// TIA Portal project "NX_PLC_Project" (V16)

(* hardware
DEVICE "S71500/ET200MP station_1"  S7-1500 station
   slot 0: "Rail_0"  Rack  6ES7 590-1***0-0AA0
   slot 0: "PM 190W 120/230VAC"  PM 190W 120/230VAC  6EP1333-4BA00
   slot 1: "PLC_1"  CPU 1516-3 PN/DP  6ES7 516-3AN01-0AB0  V2.8
      slot 3: "CPU display_1"  6ES7591-1BA00-0AA0
      slot 32768: "PROFINET interface_1"  X1
         slot 32769: "Port_1"  X1 P1
         slot 32770: "Port_2"  X1 P2
      slot 33024: "PROFINET interface_2"  X2
         slot 33025: "Port_1"  X2 P1
      slot 33280: "DP interface_1"  X3
      slot 34817: "Virtual CP interface port_1"  Virtual CP interface port  Virtual CP interface port
   slot 2: "DI 32x24VDC HF_1"  DI 32x24VDC HF  6ES7 521-1BL00-0AB0  V2.0
   slot 3: "DQ 32x24VDC/0.5A HF_1"  DQ 32x24VDC/0.5A HF  6ES7 522-1BL01-0AB0  V1.0
DEVICE "PC station"  SIMATIC PC station
   slot 0: "PC station"  Rail  SIMATIC PC-Station  V1.0
      slot 125: "Stationmanager"  Station_Manager  V6.0.4
   slot 1: "IE general_1"  IE General  IE_CP  V8.2.0
   slot 2: "HMI_RT_1"  WinCC RT Advanced  6AV2 104-0xxxx-xxxx  16.0.0.0
      slot 33792: "Computer interface"  Host interface
DEVICE "S71500/ET200MP station_2"  S7-1500 station
   slot 0: "Rail_0"  Rack  6ES7 590-1***0-0AA0
   slot 0: "PM 190W 120/230VAC"  PM 190W 120/230VAC  6EP1333-4BA00
   slot 1: "PLC_2"  CPU 1516-3 PN/DP  6ES7 516-3AN01-0AB0  V2.8
      slot 3: "CPU display_1"  6ES7591-1BA00-0AA0
      slot 32768: "PROFINET interface_1"  X1
         slot 32769: "Port_1"  X1 P1
         slot 32770: "Port_2"  X1 P2
      slot 33024: "PROFINET interface_2"  X2
         slot 33025: "Port_1"  X2 P1
      slot 33280: "DP interface_1"  X3
      slot 34817: "Virtual CP interface port_1"  Virtual CP interface port  Virtual CP interface port
   slot 2: "DI 32x24VDC HF_1"  DI 32x24VDC HF  6ES7 521-1BL00-0AB0  V2.0
   slot 3: "DQ 32x24VDC/0.5A HF_1"  DQ 32x24VDC/0.5A HF  6ES7 522-1BL01-0AB0  V1.0
DEVICE "HMI_1"  KTP700 Basic PN
   slot 0: "HMI_1"  KTP700 Basic PN  6AV2 123-2GB03-0AX0  16.0.0.0
   slot 1: "HMI_RT_2"  KTP700 Basic PN  6AV2 123-2GB03-0AX0  16.0.0.0
   slot 5: "HMI_1.IE_CP_1"  PROFINET Interface  16.0.0.0
      slot 1: "PROFINET Interface_1"  PROFINET Interface
         slot 1: "Port_1"  Port
*)

// ===== PLC "PLC_1"  CPU 1516-3 PN/DP =====

VAR_GLOBAL   // PLC tag table "Default tag table"
   "sensor1" AT %I0.0 : Bool;
   "belt1" AT %Q2.0 : Bool;
   "ABB1_ON" AT %M1.3 : Bool;
   "sensor2" AT %I0.1 : Bool;
   "sensor3" AT %I0.3 : Bool;
   "sensor4" AT %I0.4 : Bool;
   "belt2_1" AT %Q0.1 : Bool;
   "belt2_2" AT %Q0.2 : Bool;
   "belt2_3" AT %Q0.3 : Bool;
   "belt3" AT %Q0.4 : Bool;
   "send_small" AT %Q1.1 : Bool;
   "sensor2_tall" AT %I0.2 : Bool;
   "ABB2_IDLE" AT %M1.4 : Bool;
   "send_tall" AT %Q1.0 : Bool;
   "ABB2_ON" AT %M1.5 : Bool;
   "F_IDLE" AT %M0.0 : Bool;
   "FILL_TIMER_COUNT" AT %MD2 : Time;
   "ABB1_IDLE" AT %M1.2 : Bool;
   "F_SEND" AT %M0.1 : Bool;
   "robot1_end" AT %I1.1 : Bool;
   "sensor4_tall" AT %I0.5 : Bool;
   "new_cap" AT %Q1.2 : Bool;
   "F_FILL" AT %M0.2 : Bool;
   "sensor5" AT %I0.6 : Bool;
   "sensor5_tall" AT %I0.7 : Bool;
   "robot1_place_tall" AT %Q1.4 : Bool;
   "robot2_get_tall" AT %Q1.6 : Bool;
   "robot1_place_short" AT %Q1.5 : Bool;
   "robot2_get_short" AT %Q1.7 : Bool;
   "robot2_end" AT %I1.2 : Bool;
   "belt_F" AT %Q0.5 : Bool;
   "belt_L" AT %Q0.6 : Bool;
   "belt_R" AT %Q0.7 : Bool;
   "robot1_getCap" AT %Q1.3 : Bool;
   "Connect" AT %M2.0 : Bool;
   "Send" AT %M2.1 : Bool;
   "Clock_10Hz" AT %M100.0 : Bool;
   "sensor_T" AT %I2.1 : Bool;
   "ABB1_MODE" AT %M1.6 : Bool;
   "ABB2_MODE" AT %M1.7 : Bool;
   "sensor_S" AT %I2.2 : Bool;
   "ABB1_SEND" AT %M6.0 : Bool;
   "robot1_hasCap" AT %I1.0 : Bool;
   "SB_WAIT" AT %M0.3 : Bool;
   "SB_SEND" AT %M0.4 : Bool;
   "CONTROL_ENABLE" AT %M0.5 : Bool;
   "F_RELEASE" AT %M0.6 : Bool;
   "START" AT %I100.0 : Bool;
   "STOP" AT %I100.1 : Bool;
   "RESET" AT %I100.2 : Bool;
   "sink" AT %Q100.3 : Bool;
   "RESTARTING" AT %M0.7 : Bool;
   "ABB1_GETCAP" AT %M1.0 : Bool;
   "END_RESTART" AT %M1.1 : Bool;
END_VAR

DATA_BLOCK "Data_block_1"   // DB3
{ S7_Optimized_Access := 'TRUE' }
VERSION : 0.1
   VAR
      Received_string : String;
      Sent_string : String := 'Hello PLC2';
      Received_array : Array[0..1] of Char;
      Sent_array : Array[0..1] of Char;
   END_VAR
BEGIN
END_DATA_BLOCK

// folder: System blocks/Program resources

DATA_BLOCK "FILL_TIMER"   // DB1
{ S7_Optimized_Access := 'TRUE' }
AUTHOR : Simatic
FAMILY : IEC
NAME : IEC_TMR
VERSION : 1.0
// stored: InstanceOfName IEC_TIMER
"IEC_TIMER"
BEGIN
END_DATA_BLOCK

DATA_BLOCK "sink_timer"   // DB4
{ S7_Optimized_Access := 'TRUE' }
AUTHOR : Simatic
FAMILY : IEC
NAME : IEC_TMR
VERSION : 1.0
// stored: InstanceOfName IEC_TIMER
"IEC_TIMER"
BEGIN
END_DATA_BLOCK

DATA_BLOCK "PLC_1_Connection_DB"   // DB5
{ S7_Optimized_Access := 'TRUE' }
AUTHOR : SIMATIC
FAMILY : MC7Plus
NAME : TC_IP_v4
VERSION : 1.0
// stored: InstanceOfName TCON_IP_v4
"TCON_IP_v4"
BEGIN
   ID := 1;
   InterfaceId := 64;
   LocalPort := 2000;
   RemoteAddress.ADDR[1] := 192;
   RemoteAddress.ADDR[2] := 168;
   RemoteAddress.ADDR[4] := 2;
END_DATA_BLOCK

// folder: (top level)

ORGANIZATION_BLOCK "Main"   // OB1, LAD, ProgramCycle
TITLE = LADDER CODE FOR NX SIMULATION OF WATER BOTTLE ASSEMBLY LINE
{ S7_Optimized_Access := 'TRUE' }
VERSION : 0.1
// This program provides the control logic for an NX simulation via TIA Portal and PLCSIM. The simulation emulates a streamlined factory bottling line where bottles are filled, capped, and sorted for packing based on their size. The production line is organized into two primary stations:
// 
// STATION 1: Filling and Capping. This station processes the initial bottle, which is introduced from an external source (triggered via the HMI). The process begins with filling, where the bottle is conveyed to a valve and held in place for a simulated duration. Once filled, the bottle advances to the working area of ABB Robot 1. Upon detecting the bottle, the robot applies a cap and releases it toward the next stage of the line.
// 
// STATION 2: Sorting and Packing. The second station is responsible for sorting bottles by size to ensure they are packed correctly. When a bottle enters the workspace of ABB Robot 2, the robot identifies its dimensions and, following instructions from the PLC, transfers it to the appropriate secondary conveyor. Finally, the bottle travels down the designated belt to its corresponding packing crate.
// 
// IMPORTANT: The PLC program is architected using three distinct Finite State Machines (FSMs). This modular approach ensures that the Filling, Capping, and Sorting sequences operate independently yet in perfect synchronization. Without this modularity, if we used a single FSM, then instead of having mulltiple bottles going through the process, we would just be tracking a single bottle at a time and this is extremely inefficient. Having this modular approach allows us to only care about the bottles that are going through each process, not the ones moving through the belt.
// 
// IMPORTANT: Even though there are three distinct FSMs, they are connected by the sensors and the input received from the PLC's HMI, which allows us to Start, Stop, and Reset the process at any time. (We can also track the states of the robots and belts)
   VAR_INPUT
      Initial_Call : Bool;   // Initial call of this OB
      Remanence : Bool;   // =True, if remanent data are available
   END_VAR
   VAR_TEMP
      COUNT1 : Int;
      SEND_TIMER_COUNT : Time;
      cnt : UInt;
   END_VAR
   VAR_TEMP   // added for the SCL form of the ladder/FBD networks
      _w1 : Bool;
      _w2 : Bool;
      _w3 : Bool;
      _w4 : Bool;
      _w5 : Bool;
   END_VAR
BEGIN

REGION Network 1: START AND STOP LOGIC
   // This network corresponds to the START and STOP buttons in the HMI. The logic is simple: 
   // 
   // - Branch 1: If the START button is pressed, then the system (CONTROL_ENABLE) is activated.
   // 
   // - Branch 2: If the STOP button is pressed, then the system is turned off.
   // 
   // - Branch 3: If the system (CONTROL_ENABLE) is on, then belt 2 is active (belt 2 is composed of three small belts due to curving)
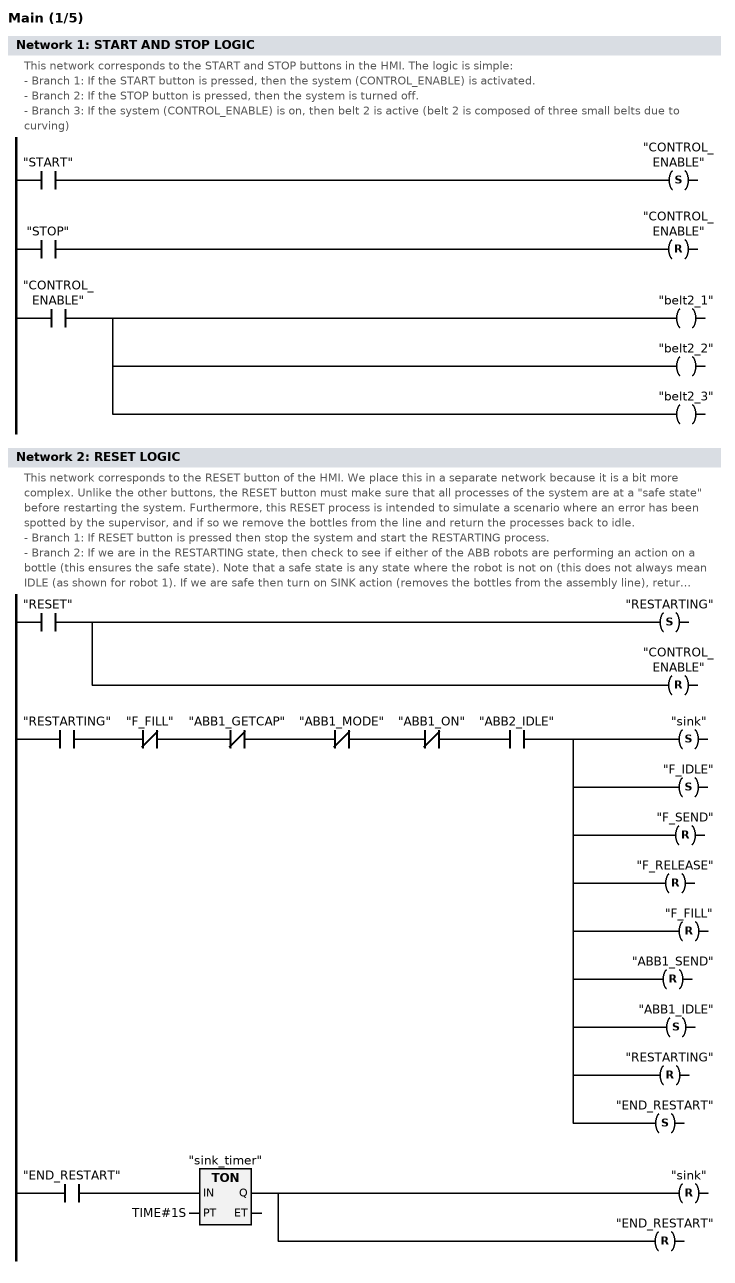
   RUNG wire#powerrail
      Contact( "START" )
      S_Coil( "CONTROL_ENABLE" )
   END_RUNG
   RUNG wire#powerrail
      Contact( "STOP" )
      R_Coil( "CONTROL_ENABLE" )
   END_RUNG
   RUNG wire#powerrail
      Contact( "CONTROL_ENABLE" )
      wire#w1
      Coil( "belt2_1" )
   END_RUNG
   RUNG wire#w1
      Coil( "belt2_2" )
   END_RUNG
   RUNG wire#w1
      Coil( "belt2_3" )
   END_RUNG
   // the same network as SCL:
   IF "START" THEN "CONTROL_ENABLE" := TRUE; END_IF;
   IF "STOP" THEN "CONTROL_ENABLE" := FALSE; END_IF;
   "belt2_1" := "CONTROL_ENABLE";
   "belt2_2" := "CONTROL_ENABLE";
   "belt2_3" := "CONTROL_ENABLE";
END_REGION

REGION Network 2: RESET LOGIC
   // This network corresponds to the RESET button of the HMI. We place this in a separate network because it is a bit more complex. Unlike the other buttons, the RESET button must make sure that all processes of the system are at a "safe state" before restarting the system. Furthermore, this RESET process is intended to simulate a scenario where an error has been spotted by the supervisor, and if so we remove the bottles from the line and return the processes back to idle. 
   // 
   // - Branch 1: If RESET button is pressed then stop the system and start the RESTARTING process.
   // 
   // - Branch 2: If we are in the RESTARTING state, then check to see if either of the ABB robots are performing an action on a bottle (this ensures the safe state). Note that a safe state is any state where the robot is not on (this does not always mean IDLE (as shown for robot 1). If we are safe then turn on SINK action (removes the bottles from the assembly line), return FSMs to Idle and move to END_RESTART state. Note that we only reset the states that can possibly be active (some states we know for sure are off).
   // 
   // - Branch 3: This END_RESTART state is made to ensure the sinking action is performed because using a single coil gives errors due to NX synchronization. In a perfect scenario using a single coil in the previous branched would have sufficed.
   // 
   // After resetting, the user must again press START, as well as send a new bottle and place a new cap for ABB robot 1.
   IF "RESET" THEN
       "RESTARTING" := TRUE;
       "CONTROL_ENABLE" := FALSE;
   END_IF;
   IF "RESTARTING" AND NOT "F_FILL" AND NOT "ABB1_GETCAP" AND NOT "ABB1_MODE" AND NOT "ABB1_ON" AND "ABB2_IDLE" THEN
       "sink" := TRUE;
       "F_IDLE" := TRUE;
       "F_SEND" := FALSE;
       "F_RELEASE" := FALSE;
   END_IF;
   #_w1 := "RESTARTING" AND NOT "F_FILL" AND NOT "ABB1_GETCAP" AND NOT "ABB1_MODE" AND NOT "ABB1_ON" AND "ABB2_IDLE";
   IF #_w1 THEN
       "F_FILL" := FALSE;
       "ABB1_SEND" := FALSE;
       "ABB1_IDLE" := TRUE;
       "RESTARTING" := FALSE;
       "END_RESTART" := TRUE;
   END_IF;
   "sink_timer".TON(IN := "END_RESTART", PT := TIME#1S);
   IF "sink_timer".Q THEN
       "sink" := FALSE;
       "END_RESTART" := FALSE;
   END_IF;
END_REGION

REGION Network 3: FILLING PROCESS
   // This station corresponds to the filling process in station 1. Here the bottle starts at the beggining of belt1, moves to the valve, is filled, and sent along to the next process.
   // 
   // - Branch 1: Initial scenario, IDLE is the first state of this FSM.
   // 
   // - Branch 2: If IDLE and system is on, and either of the sensors detect a bottle at the top of belt 1, then move to SEND state.
   // 
   // - Branch 3: This SEND state checks if the system is on, and when the bottle reaches sensor 1, we move to the FILL state. Note that the belt is moving during this, it is done in the last branch of this network.
   // 
   // - Branch 4: The FILL state checks if  sensor 1 is activate. If so we start a timer to simulate filling. Once the timer hits, we move on to the RELEASE state. Note that this state does not check if the system is enabled, this is to ensure that the filling process finishes if the restart button is pressed (safe state).
   // 
   // - Branch 5: During this RELEASE state, belt 1 is moving and we are checking if the bottle reaches sensor 2, if so then this means the bottle has left belt 1 and is now at belt 2. Finally we move back to IDLE.
   // 
   // - Branch 6: If we are at states SEND or RELEASE and the system is active, then we move belt 1.
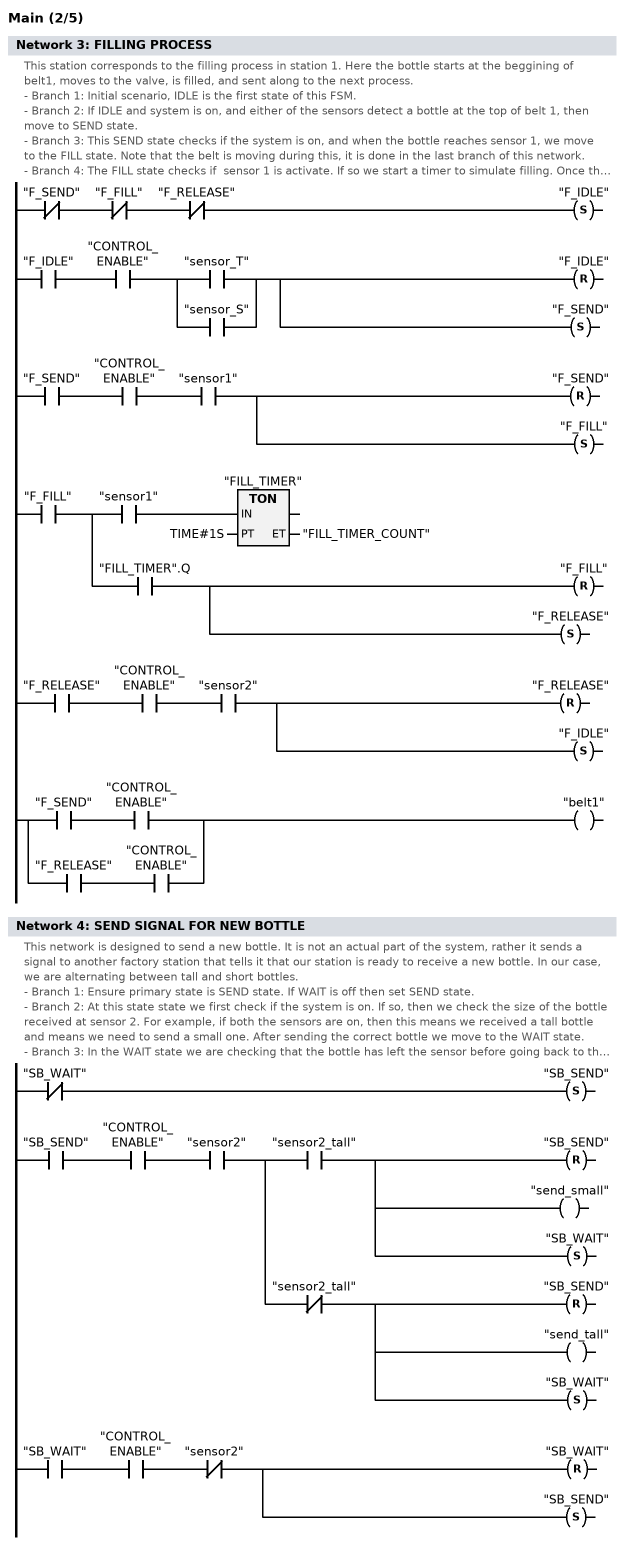
   IF NOT "F_SEND" AND NOT "F_FILL" AND NOT "F_RELEASE" THEN "F_IDLE" := TRUE; END_IF;
   #_w1 := "F_IDLE" AND "CONTROL_ENABLE" AND ("sensor_T" OR "sensor_S");
   IF #_w1 THEN
       "F_IDLE" := FALSE;
       "F_SEND" := TRUE;
   END_IF;
   #_w2 := "F_SEND" AND "CONTROL_ENABLE" AND "sensor1";
   IF #_w2 THEN
       "F_SEND" := FALSE;
       "F_FILL" := TRUE;
   END_IF;
   "FILL_TIMER".TON(IN := "F_FILL" AND "sensor1", PT := TIME#1S, ET => "FILL_TIMER_COUNT");
   #_w3 := "F_FILL" AND "FILL_TIMER".Q;
   IF #_w3 THEN
       "F_FILL" := FALSE;
       "F_RELEASE" := TRUE;
   END_IF;
   #_w4 := "F_RELEASE" AND "CONTROL_ENABLE" AND "sensor2";
   IF #_w4 THEN
       "F_RELEASE" := FALSE;
       "F_IDLE" := TRUE;
   END_IF;
   "belt1" := ("F_SEND" AND "CONTROL_ENABLE") OR ("F_RELEASE" AND "CONTROL_ENABLE");
END_REGION

REGION Network 4: SEND SIGNAL FOR NEW BOTTLE
   // This network is designed to send a new bottle. It is not an actual part of the system, rather it sends a signal to another factory station that tells it that our station is ready to receive a new bottle. In our case, we are alternating between tall and short bottles.
   // 
   // - Branch 1: Ensure primary state is SEND state. If WAIT is off then set SEND state.
   // 
   // - Branch 2: At this state state we first check if the system is on. If so, then we check the size of the bottle received at sensor 2. For example, if both the sensors are on, then this means we received a tall bottle and means we need to send a small one. After sending the correct bottle we move to the WAIT state.
   // 
   // - Branch 3: In the WAIT state we are checking that the bottle has left the sensor before going back to the SEND state. This is necessary, without it the system would send multiple bottles.
   RUNG wire#powerrail
      I_Contact( "SB_WAIT" )
      S_Coil( "SB_SEND" )
   END_RUNG
   RUNG wire#powerrail
      Contact( "SB_SEND" )
      Contact( "CONTROL_ENABLE" )
      Contact( "sensor2" )
      wire#w1
      Contact( "sensor2_tall" )
      wire#w2
      R_Coil( "SB_SEND" )
   END_RUNG
   RUNG wire#w2
      Coil( "send_small" )
   END_RUNG
   RUNG wire#w2
      S_Coil( "SB_WAIT" )
   END_RUNG
   RUNG wire#w1
      I_Contact( "sensor2_tall" )
      wire#w3
      R_Coil( "SB_SEND" )
   END_RUNG
   RUNG wire#w3
      Coil( "send_tall" )
   END_RUNG
   RUNG wire#w3
      S_Coil( "SB_WAIT" )
   END_RUNG
   RUNG wire#powerrail
      Contact( "SB_WAIT" )
      Contact( "CONTROL_ENABLE" )
      I_Contact( "sensor2" )
      wire#w4
      R_Coil( "SB_WAIT" )
   END_RUNG
   RUNG wire#w4
      S_Coil( "SB_SEND" )
   END_RUNG
   // the same network as SCL:
   IF NOT "SB_WAIT" THEN "SB_SEND" := TRUE; END_IF;
   #_w1 := "SB_SEND" AND "CONTROL_ENABLE" AND "sensor2";
   #_w2 := #_w1 AND "sensor2_tall";
   IF #_w2 THEN "SB_SEND" := FALSE; END_IF;
   "send_small" := #_w2;
   IF #_w2 THEN "SB_WAIT" := TRUE; END_IF;
   #_w3 := #_w1 AND NOT "sensor2_tall";
   IF #_w3 THEN "SB_SEND" := FALSE; END_IF;
   "send_tall" := #_w3;
   IF #_w3 THEN "SB_WAIT" := TRUE; END_IF;
   #_w4 := "SB_WAIT" AND "CONTROL_ENABLE" AND NOT "sensor2";
   IF #_w4 THEN
       "SB_WAIT" := FALSE;
       "SB_SEND" := TRUE;
   END_IF;
END_REGION

REGION Network 5: ABB ROBOT 1 - CAPPING PROCESS
   // This network corresponds to the FSM for the capping process performed by ABB Robot 1. Here the bottle reaches the sensor in the robot's workspace and starts the process. Note that the states in branches 3, 4, and 5, do not check if the system is on, this is crucial to ensure that the robot finishes the current operation before stopping (safe state).
   // 
   // - Branch 1: Initial scenario of this FSM. IDLE is the first state.
   // 
   // - Branch 2: At IDLE state we check if the system is on, as well as if the bottle has reached the robot's sensor. If so then send a signal to the robot to get the cap and move to GETCAP state.
   // 
   // - Branch 3: The GETCAP state checks for a confirmation signal from the robot (in NX) to ensure the robot has the cap and is in position. If so we reset the signal and move to the MODE state. 
   // 
   // - Branch 4: The MODE state is similar to the "send_bottle" process, where we check the size of the bottle. Once checked, we send the correct signal to the robot (either tall or short placing). We then move to the ON state.
   // 
   // - Branch 5: The ON state checks for confirmation from the robot that it has finished the placing action. If so we create a new cap and reset the placing signals of the robot. We then move to the SEND state.
   // 
   // - Branch 6: The SEND state works similarly to the "wait state" in the send bottle process, we wait until the bottle passes the sensor before returning to the IDLE state. This ensures the robot does not mistake it for a new bottle. FInally we move back to IDLE.
   // 
   // - Branch 7: If system is active and we are at IDLE or SEND, then we activate belt 3.
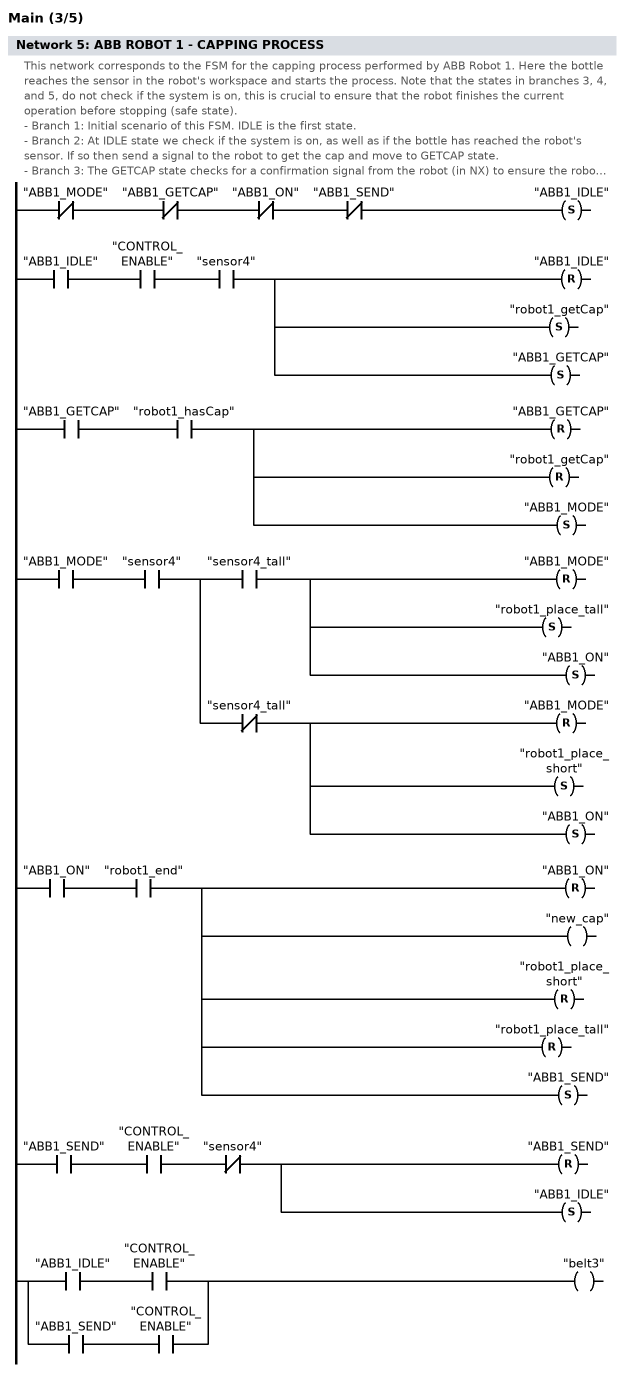
   RUNG wire#powerrail
      I_Contact( "ABB1_MODE" )
      I_Contact( "ABB1_GETCAP" )
      I_Contact( "ABB1_ON" )
      I_Contact( "ABB1_SEND" )
      S_Coil( "ABB1_IDLE" )
   END_RUNG
   RUNG wire#powerrail
      Contact( "ABB1_IDLE" )
      Contact( "CONTROL_ENABLE" )
      Contact( "sensor4" )
      wire#w1
      R_Coil( "ABB1_IDLE" )
   END_RUNG
   RUNG wire#w1
      S_Coil( "robot1_getCap" )
   END_RUNG
   RUNG wire#w1
      S_Coil( "ABB1_GETCAP" )
   END_RUNG
   RUNG wire#powerrail
      Contact( "ABB1_GETCAP" )
      Contact( "robot1_hasCap" )
      wire#w2
      R_Coil( "ABB1_GETCAP" )
   END_RUNG
   RUNG wire#w2
      R_Coil( "robot1_getCap" )
   END_RUNG
   RUNG wire#w2
      S_Coil( "ABB1_MODE" )
   END_RUNG
   RUNG wire#powerrail
      Contact( "ABB1_MODE" )
      Contact( "sensor4" )
      wire#w3
      Contact( "sensor4_tall" )
      wire#w4
      R_Coil( "ABB1_MODE" )
   END_RUNG
   RUNG wire#w4
      S_Coil( "robot1_place_tall" )
   END_RUNG
   RUNG wire#w4
      S_Coil( "ABB1_ON" )
   END_RUNG
   RUNG wire#w3
      I_Contact( "sensor4_tall" )
      wire#w5
      R_Coil( "ABB1_MODE" )
   END_RUNG
   RUNG wire#w5
      S_Coil( "robot1_place_short" )
   END_RUNG
   RUNG wire#w5
      S_Coil( "ABB1_ON" )
   END_RUNG
   RUNG wire#powerrail
      Contact( "ABB1_ON" )
      Contact( "robot1_end" )
      wire#w6
      R_Coil( "ABB1_ON" )
   END_RUNG
   RUNG wire#w6
      Coil( "new_cap" )
   END_RUNG
   RUNG wire#w6
      R_Coil( "robot1_place_short" )
   END_RUNG
   RUNG wire#w6
      R_Coil( "robot1_place_tall" )
   END_RUNG
   RUNG wire#w6
      S_Coil( "ABB1_SEND" )
   END_RUNG
   RUNG wire#powerrail
      Contact( "ABB1_SEND" )
      Contact( "CONTROL_ENABLE" )
      I_Contact( "sensor4" )
      wire#w7
      R_Coil( "ABB1_SEND" )
   END_RUNG
   RUNG wire#w7
      S_Coil( "ABB1_IDLE" )
   END_RUNG
   RUNG wire#powerrail
      Contact( "ABB1_IDLE" )
      Contact( "CONTROL_ENABLE" )
      wire#w8
      Coil( "belt3" )
   END_RUNG
   RUNG wire#powerrail
      Contact( "ABB1_SEND" )
      Contact( "CONTROL_ENABLE" )
   END_RUNG wire#w8
   // the same network as SCL:
   IF NOT "ABB1_MODE" AND NOT "ABB1_GETCAP" AND NOT "ABB1_ON" AND NOT "ABB1_SEND" THEN
       "ABB1_IDLE" := TRUE;
   END_IF;
   #_w1 := "ABB1_IDLE" AND "CONTROL_ENABLE" AND "sensor4";
   IF #_w1 THEN
       "ABB1_IDLE" := FALSE;
       "robot1_getCap" := TRUE;
       "ABB1_GETCAP" := TRUE;
   END_IF;
   #_w2 := "ABB1_GETCAP" AND "robot1_hasCap";
   IF #_w2 THEN
       "ABB1_GETCAP" := FALSE;
       "robot1_getCap" := FALSE;
       "ABB1_MODE" := TRUE;
   END_IF;
   #_w3 := "ABB1_MODE" AND "sensor4";
   IF #_w3 AND "sensor4_tall" THEN
       "ABB1_MODE" := FALSE;
       "robot1_place_tall" := TRUE;
       "ABB1_ON" := TRUE;
   END_IF;
   IF #_w3 AND NOT "sensor4_tall" THEN
       "ABB1_MODE" := FALSE;
       "robot1_place_short" := TRUE;
       "ABB1_ON" := TRUE;
   END_IF;
   #_w4 := "ABB1_ON" AND "robot1_end";
   IF #_w4 THEN "ABB1_ON" := FALSE; END_IF;
   "new_cap" := #_w4;
   IF #_w4 THEN
       "robot1_place_short" := FALSE;
       "robot1_place_tall" := FALSE;
       "ABB1_SEND" := TRUE;
   END_IF;
   #_w5 := "ABB1_SEND" AND "CONTROL_ENABLE" AND NOT "sensor4";
   IF #_w5 THEN
       "ABB1_SEND" := FALSE;
       "ABB1_IDLE" := TRUE;
   END_IF;
   "belt3" := ("ABB1_IDLE" AND "CONTROL_ENABLE") OR ("ABB1_SEND" AND "CONTROL_ENABLE");
END_REGION

REGION Network 6: ABB ROBOT 2 - SORTING PROCESS
   // This network corresponds to the FSM for ABB Robot 2. This is the process of sorting bottles and placing them in the correct conveyor belt, where the bottle will move to a packing box. Note that the states in branches 3 and 4 do not check if the system is on, as explained before, this is to ensure the robot ends its current action before stopping the system.
   // 
   // - Branch 1: Initailization of FSM. IDLE is the first state.
   // 
   // - Branch 2: At IDLE state, we check if the system is active. We check if the sensor in the robot's workspace, and if so we move on to the MODE state. 
   // 
   // - Branch 3: At the MODE state, we again check the size of the bottle through the use of two sensors. We then send the corresponding signal to the robot (in the NX simulation) and move to the ON state.
   // 
   // - Branch 4: At the ON state we check for the confirmation signal from the robot. If we receive the signal this means the robot has ended the action, and therefore we reset the signals and move back to the IDLE state.
   // 
   // 
   // - Branch 5:  If system is active and we are at IDLE, then we activate belts F, L, and R.
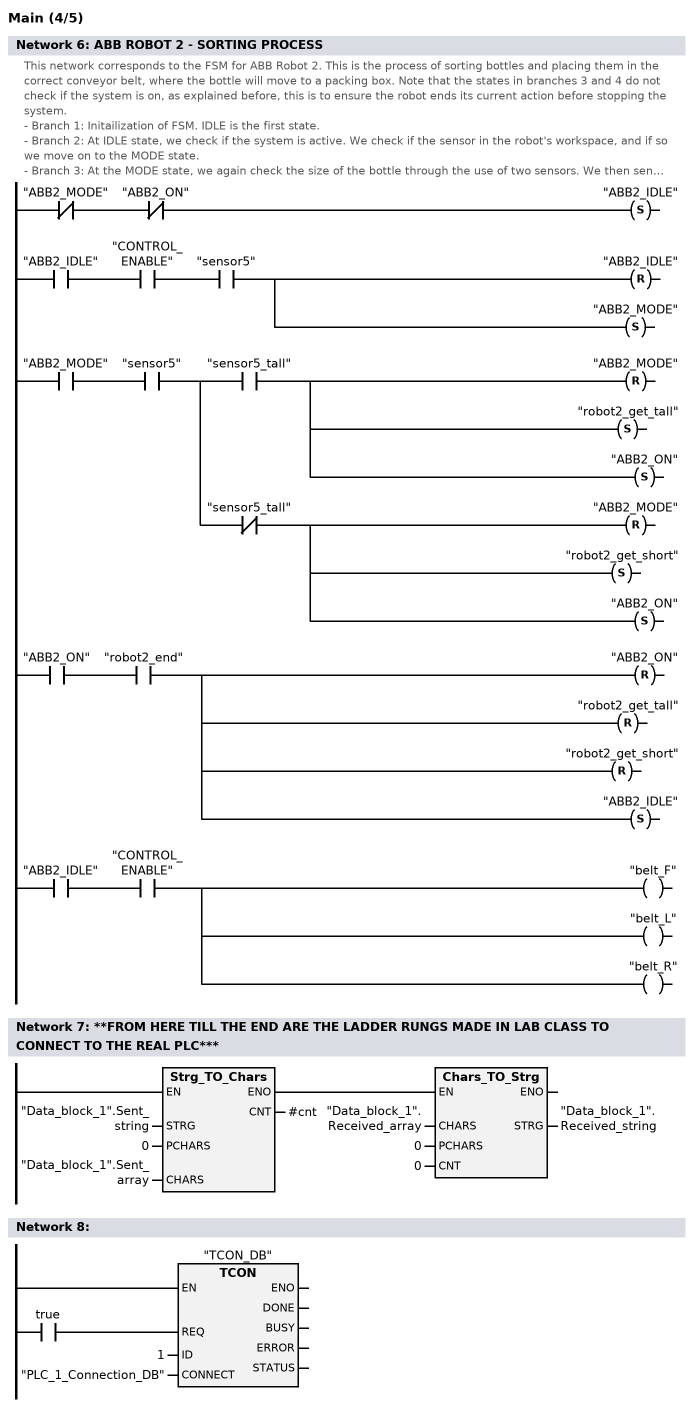
   RUNG wire#powerrail
      I_Contact( "ABB2_MODE" )
      I_Contact( "ABB2_ON" )
      S_Coil( "ABB2_IDLE" )
   END_RUNG
   RUNG wire#powerrail
      Contact( "ABB2_IDLE" )
      Contact( "CONTROL_ENABLE" )
      Contact( "sensor5" )
      wire#w1
      R_Coil( "ABB2_IDLE" )
   END_RUNG
   RUNG wire#w1
      S_Coil( "ABB2_MODE" )
   END_RUNG
   RUNG wire#powerrail
      Contact( "ABB2_MODE" )
      Contact( "sensor5" )
      wire#w2
      Contact( "sensor5_tall" )
      wire#w3
      R_Coil( "ABB2_MODE" )
   END_RUNG
   RUNG wire#w3
      S_Coil( "robot2_get_tall" )
   END_RUNG
   RUNG wire#w3
      S_Coil( "ABB2_ON" )
   END_RUNG
   RUNG wire#w2
      I_Contact( "sensor5_tall" )
      wire#w4
      R_Coil( "ABB2_MODE" )
   END_RUNG
   RUNG wire#w4
      S_Coil( "robot2_get_short" )
   END_RUNG
   RUNG wire#w4
      S_Coil( "ABB2_ON" )
   END_RUNG
   RUNG wire#powerrail
      Contact( "ABB2_ON" )
      Contact( "robot2_end" )
      wire#w5
      R_Coil( "ABB2_ON" )
   END_RUNG
   RUNG wire#w5
      R_Coil( "robot2_get_tall" )
   END_RUNG
   RUNG wire#w5
      R_Coil( "robot2_get_short" )
   END_RUNG
   RUNG wire#w5
      S_Coil( "ABB2_IDLE" )
   END_RUNG
   RUNG wire#powerrail
      Contact( "ABB2_IDLE" )
      Contact( "CONTROL_ENABLE" )
      wire#w6
      Coil( "belt_F" )
   END_RUNG
   RUNG wire#w6
      Coil( "belt_L" )
   END_RUNG
   RUNG wire#w6
      Coil( "belt_R" )
   END_RUNG
   // the same network as SCL:
   IF NOT "ABB2_MODE" AND NOT "ABB2_ON" THEN "ABB2_IDLE" := TRUE; END_IF;
   #_w1 := "ABB2_IDLE" AND "CONTROL_ENABLE" AND "sensor5";
   IF #_w1 THEN
       "ABB2_IDLE" := FALSE;
       "ABB2_MODE" := TRUE;
   END_IF;
   #_w2 := "ABB2_MODE" AND "sensor5";
   IF #_w2 AND "sensor5_tall" THEN
       "ABB2_MODE" := FALSE;
       "robot2_get_tall" := TRUE;
       "ABB2_ON" := TRUE;
   END_IF;
   IF #_w2 AND NOT "sensor5_tall" THEN
       "ABB2_MODE" := FALSE;
       "robot2_get_short" := TRUE;
       "ABB2_ON" := TRUE;
   END_IF;
   #_w3 := "ABB2_ON" AND "robot2_end";
   IF #_w3 THEN
       "ABB2_ON" := FALSE;
       "robot2_get_tall" := FALSE;
       "robot2_get_short" := FALSE;
       "ABB2_IDLE" := TRUE;
   END_IF;
   "belt_F" := "ABB2_IDLE" AND "CONTROL_ENABLE";
   "belt_L" := "belt_F";
   "belt_R" := "belt_F";
END_REGION

REGION Network 7: **FROM HERE TILL THE END ARE THE LADDER RUNGS MADE IN LAB CLASS TO CONNECT TO THE REAL PLC***
   // no SCL statement known for Chars_TO_Strg, Strg_TO_Chars: written as a call
   // ENO of a box is taken as its EN; it also drops when the box reports an error
   Strg_TO_Chars(Strg := "Data_block_1".Sent_string,
                 pChars := 0,
                 Chars := "Data_block_1".Sent_array,
                 Cnt => #cnt);
   Chars_TO_Strg(Chars := "Data_block_1".Received_array,
                 pChars := 0,
                 Cnt := 0,
                 Strg => "Data_block_1".Received_string);
END_REGION

REGION Network 8
   "TCON_DB"(REQ := true, ID := 1, CONNECT := "PLC_1_Connection_DB");   // TCON
END_REGION

REGION Network 9
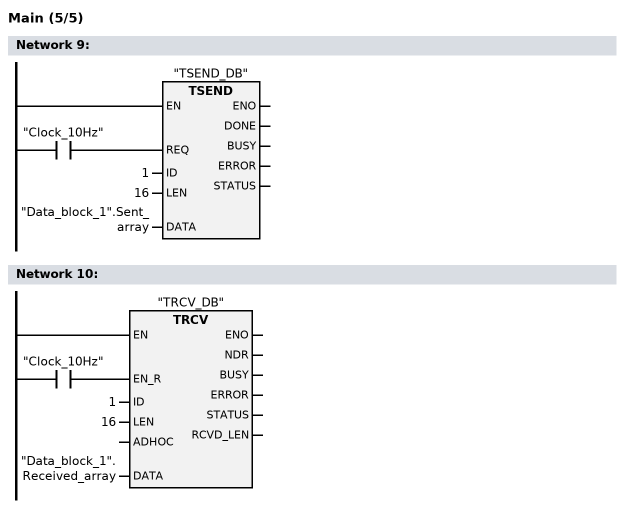
   "TSEND_DB"(REQ := "Clock_10Hz", ID := 1, LEN := 16, DATA := "Data_block_1".Sent_array);   // TSEND
END_REGION

REGION Network 10
   "TRCV_DB"(EN_R := "Clock_10Hz", ID := 1, LEN := 16, DATA := "Data_block_1".Received_array);   // TRCV
END_REGION
END_ORGANIZATION_BLOCK

// ===== PLC "PLC_2"  CPU 1516-3 PN/DP =====

VAR_GLOBAL   // PLC tag table "PLC2_tag_table"
   "sensor1" AT %I0.0 : Bool;   // INPUT FOR SENSOR 1 --> FOR FILLING
   "sensor2" AT %I0.1 : Bool;   // INPUT FOR SENSOR 2 --> FOR OBJ SOURCE CREATION
   "sensor2_tall" AT %I0.2 : Bool;   // INPUT FOR SENSOR 2 TALL --> FOR OBJ SOURCE CREATION
   "sensor3" AT %I0.3 : Bool;   // INPUT FOR SENSOR 3 --> FOR CONTROLLING THE FLOW OF THE BOTTLES
   "sensor4" AT %I0.4 : Bool;   // INPUT FOR SENSOR 4 --> FOR ROBOT 1 OPERATIONS
   "sensor4_tall" AT %I0.5 : Bool;   // INPUT FOR SENSOR 4 TALL --> FOR ROBOT 1 OPERATIONS
   "sensor5" AT %I0.6 : Bool;   // INPUT FOR SENSOR 5 --> FOR ROBOT 2 OPERATIONS
   "sensor5_tall" AT %I0.7 : Bool;   // INPUT FOR SENSOR 5 TALL --> FOR ROBOT 2 OPERATIONS
   "robot1_end" AT %I1.1 : Bool;   // INPUT FOR ROBOT1_END --> FOR SIGNALING END OF ROBOT 1 OPERATIONS
   "robot2_end" AT %I1.2 : Bool;   // INPUT FOR ROBOT2_END --> FOR SIGNALING END OF ROBOT 2 OPERATIONS
   "belt1" AT %Q0.0 : Bool;   // OUTPUT FOR BELT 1 --> TURN ON/OFF CONVEYOR BELT 1
   "belt2_1" AT %Q0.1 : Bool;   // OUTPUT FOR BELT 2.1 --> TURN ON/OFF CONVEYOR BELT 2.1
   "belt2_2" AT %Q0.2 : Bool;   // OUTPUT FOR BELT 2.2 --> TURN ON/OFF CONVEYOR BELT 2.2
   "belt2_3" AT %Q0.3 : Bool;   // OUTPUT FOR BELT 2.3 --> TURN ON/OFF CONVEYOR BELT 2.3
   "belt3" AT %Q0.4 : Bool;   // OUTPUT FOR BELT 3 --> TURN ON/OFF CONVEYOR BELT 3
   "belt_F" AT %Q0.5 : Bool;   // OUTPUT FOR BELT F --> TURN ON/OFF CONVEYOR BELT F (IN FRONT OF ROBOT 2)
   "belt_L" AT %Q0.6 : Bool;   // OUTPUT FOR BELT L --> TURN ON/OFF CONVEYOR BELT L (LEFT OF ROBOT 2)
   "belt_R" AT %Q0.7 : Bool;   // OUTPUT FOR BELT R --> TURN ON/OFF CONVEYOR BELT R (RIGHT OF ROBOT 2)
   "send_tall" AT %Q1.0 : Bool;   // OUTPUT FOR SEND_TALL --> FOR SENDING A NEW TALL BOTTLE
   "send_small" AT %Q1.1 : Bool;   // OUTPUT FOR SEND_SMALL --> FOR SENDING A NEW SMALL BOTTLE
   "new_cap" AT %Q1.2 : Bool;   // OUTPUT FOR NEW_CAP --> FOR SENDING A NEW CAP
   "robot1_getCap" AT %Q1.3 : Bool;   // OUTPUT FOR ROBOT1_GETCAP --> TELLS ROBOT 1 TO GET CAP FROM BOX
   "robot1_place_tall" AT %Q1.4 : Bool;   // OUTPUT FOR ROBOT1_PLACETALL --> TELLS ROBOT 1 TO PERFORM SEQUENCE FOR TALL
   "robot1_place_short" AT %Q1.5 : Bool;   // OUTPUT FOR ROBOT1_PLACESHORT --> TELLS ROBOT 1 TO PERFORM SEQUENCE FOR SHORT
   "robot2_get_tall" AT %Q1.6 : Bool;   // OUTPUT FOR ROBOT2_PLACETALL --> TELLS ROBOT 2 TO PERFORM SEQUENCE FOR TALL
   "robot2_get_short" AT %Q1.7 : Bool;   // OUTPUT FOR ROBOT2_PLACESHORT --> TELLS ROBOT 2 TO PERFORM SEQUENCE FOR SHORT
   "START" AT %M0.0 : Bool;   // STATE FOR START --> INITIALIZATION STATE
   "ROBOT_STATION1" AT %M0.1 : Bool;   // STATE FOR ROBOT_STATION1 --> LOGIC FOR ROBOT 1
   "ROBOT_STATION2" AT %M0.2 : Bool;   // STATE FOR ROBOT_STATION2 --> LOGIC FOR ROBOT 2
   "SEND_TO_FILL" AT %M1.0 : Bool;   // STATE FOR SEND_TO_FILL --> FOR SENDING BOTTLE TO FILLER
   "FILL" AT %M1.1 : Bool;   // STATE FOR FILL --> FOR SIMULATING THE FILLER ACTION
   "CHOOSE_NEW_BOTTLE" AT %M1.2 : Bool;   // STATE FOR CHOOSE_NEW_BOTTLE --> DECIDE WHICH BOTTLE TO SEND
   "SEND_NEW_SMALL" AT %M1.3 : Bool;   // STATE FOR SEND_NEW_SMALL --> FOR SENDING A SMALL BOTTLE
   "SEND_NEW_TALL" AT %M1.4 : Bool;   // STATE FOR SEND_NEW_TALL --> FOR SENDING A TALL BOTTLE
   "TRANSITION" AT %M1.5 : Bool;   // STATE FOR TRANSITION --> FOR CONTROLLING THE LOGIC OF THE FLOW
   "WAIT_TO_SEND" AT %M1.6 : Bool;   // STATE FOR WAIT_TO_SEND --> FOR WAITING TO SEND TO ROBOT 1
   "SEND_TO_PLACE" AT %M1.7 : Bool;   // STATE FOR SEND_TO_PLACE --> FOR SENDING BOTTLE TO ROBOT 1
   "FILL_TIMER_COUNT" AT %MD2 : Time;   // TIMER FILL_TIMER_COUNT --> 1 SECOND TIMER TO SIMULATE FILLING
   "Connect" AT %M2.0 : Bool;
   "Send" AT %M2.1 : Bool;
   "Clock_10Hz" AT %M200.0 : Bool;
   "Clock_Byte" AT %MB200 : Byte;
   "Clock_10Hz(1)" AT %M0.0 : Bool;
   "Clock_5Hz" AT %M200.1 : Bool;
   "Clock_2.5Hz" AT %M200.2 : Bool;
   "Clock_2Hz" AT %M200.3 : Bool;
   "Clock_1.25Hz" AT %M200.4 : Bool;
   "Clock_1Hz" AT %M200.5 : Bool;
   "Clock_0.625Hz" AT %M200.6 : Bool;
   "Clock_0.5Hz" AT %M200.7 : Bool;
END_VAR

DATA_BLOCK "PLC2_Data_block_1"   // DB4
{ S7_Optimized_Access := 'TRUE' }
VERSION : 0.1
   VAR
      Received_string : String;
      Sent_string : String := 'Hello PLC1';
      Received_array : Array[0..1] of Char;
      Sent_array : Array[0..1] of Char;
   END_VAR
BEGIN
END_DATA_BLOCK

// folder: System blocks/Program resources

DATA_BLOCK "PLC_2_Connection_DB"   // DB3
{ S7_Optimized_Access := 'TRUE' }
AUTHOR : SIMATIC
FAMILY : MC7Plus
NAME : TC_IP_v4
VERSION : 1.0
// stored: InstanceOfName TCON_IP_v4
"TCON_IP_v4"
BEGIN
   ID := 1;
   InterfaceId := 64;
   RemotePort := 2000;
   ActiveEstablished := true;
   RemoteAddress.ADDR[1] := 192;
   RemoteAddress.ADDR[2] := 168;
   RemoteAddress.ADDR[4] := 4;
END_DATA_BLOCK

// folder: (top level)

ORGANIZATION_BLOCK "PLC2_Main"   // OB1, LAD, ProgramCycle
TITLE = "Main Program Sweep (Cycle)"
{ S7_Optimized_Access := 'TRUE' }
VERSION : 0.1
   VAR_INPUT
      Initial_Call : Bool;   // Initial call of this OB
      Remanence : Bool;   // =True, if remanent data are available
   END_VAR
   VAR_TEMP
      COUNT1 : Int;
      SEND_TIMER_COUNT : Time;
   END_VAR
BEGIN

REGION Network 1
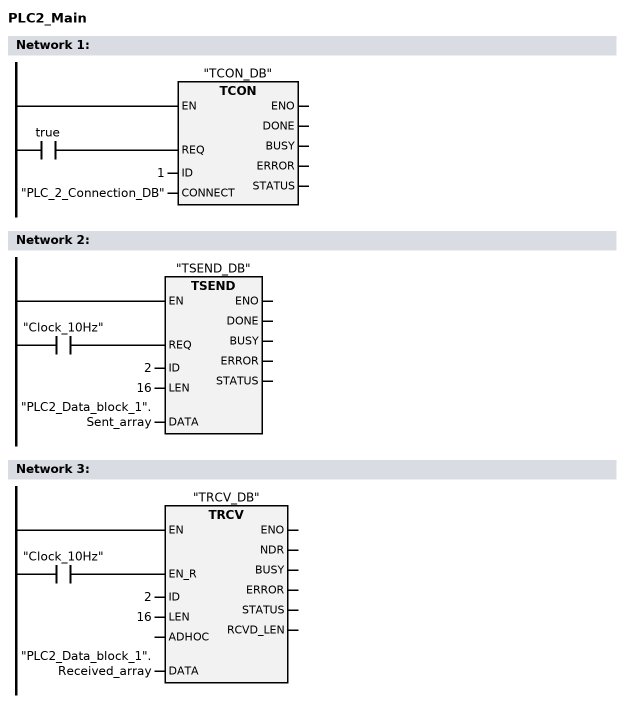
   "TCON_DB"(REQ := true, ID := 1, CONNECT := "PLC_2_Connection_DB");   // TCON
END_REGION

REGION Network 2
   "TSEND_DB"(REQ := "Clock_10Hz", ID := 2, LEN := 16, DATA := "PLC2_Data_block_1".Sent_array);   // TSEND
END_REGION

REGION Network 3
   "TRCV_DB"(EN_R := "Clock_10Hz", ID := 2, LEN := 16, DATA := "PLC2_Data_block_1".Received_array);   // TRCV
END_REGION
END_ORGANIZATION_BLOCK

(* ===== HMI "HMI_RT_1" =====
system functions are stored by id; their names below are inferred from use
connection "HMI_Connection_2": ETHERNET, S7_1500_OMS

HMI tags "Default tag table"
   "START" : Bool = PLC START AT %I100.0, 1 s

screen "Screen_1" 1024x768
   Button "Button_1" at 434,242 size 112x51; TextOff 'START'
      on Press: SetBit("START")
      on Release: ResetBit("START")
*)

(* ===== HMI "HMI_RT_2" =====
system functions are stored by id; their names below are inferred from use
connection "HMI_Connection_1": ETHERNET, SMART_S7_1500_OMS

HMI tags "Default tag table"
   "Tag_ScreenNumber" : UInt, internal
   "START" : Bool = PLC START AT %I100.0, 100 ms
   "STOP" : Bool = PLC STOP AT %I100.1, 100 ms
   "send_tall" : Bool = PLC send_tall AT %Q1.0, 100 ms
   "send_small" : Bool = PLC send_small AT %Q1.1, 100 ms
   "CONTROL_ENABLE" : Bool = PLC CONTROL_ENABLE AT %M0.5, 1 s
   "belt1" : Bool = PLC belt1 AT %Q2.0, 1 s
   "belt2_1" : Bool = PLC belt2_1 AT %Q0.1, 1 s
   "belt3" : Bool = PLC belt3 AT %Q0.4, 1 s
   "belt_F" : Bool = PLC belt_F AT %Q0.5, 1 s
   "belt_R" : Bool = PLC belt_R AT %Q0.7, 1 s
   "belt_L" : Bool = PLC belt_L AT %Q0.6, 1 s
   "ABB1_IDLE" : Bool = PLC ABB1_IDLE AT %M1.2, 1 s
   "ABB2_IDLE" : Bool = PLC ABB2_IDLE AT %M1.4, 1 s
   "RESET" : Bool = PLC RESET AT %I100.2, 1 s
   "RESTARTING" : Bool = PLC RESTARTING AT %M0.7, 1 s
   "F_FILL" : Bool = PLC F_FILL AT %M0.2, 1 s
   "new_cap" : Bool = PLC new_cap AT %Q1.2, 1 s

Template "Template_1" 800x480
   Button "Exit" at 714,429 size 71x50; TextOff 'Exit'; PictureOff "ExitRuntime_KTP700_Basic_PN_TR"; PictureOn "ExitRuntime_KTP700_Basic_PN_TR"
      on Release: StopRuntime(0)
   Button "Template_Button" at 614,429 size 71x50; TextOff 'Text'
   Button "Template_Button_1" at 514,429 size 71x50; TextOff 'Text'
   Button "Template_Button_2" at 414,429 size 71x50; TextOff 'Text'
   Button "Template_Button_3" at 314,429 size 71x50; TextOff 'Text'
   Button "Template_Button_4" at 214,429 size 71x50; TextOff 'Text'
   Button "Template_Button_5" at 114,429 size 71x50; TextOff 'Text'
   Button "Start screen" at 14,429 size 71x50; TextOff 'Start screen'; PictureOff "NavigateHome_KTP700_Basic_PN_TR"; PictureOn "NavigateHome_KTP700_Basic_PN_TR"
      on Release: ActivateScreen("Root screen", 0)
   SymbolicIOField "Symbolic_IO_Field_Screen" at 93,9 size 600x33; TextOff '0'; TextOn '1'; TextList "TextList_ScreenNames"
      ProcessValue <- "Tag_ScreenNumber"
      on Change: ActivateScreenByNumber("Tag_ScreenNumber", 0)
   DateTimeField "HmiScreenItemData" at 695,25 size 105x25
   DateTimeField "HmiScreenItemData_1" at 695,0 size 105x25
   GraphicView "Logo" at 0,0 size 91x51; Picture "Logo of HMI_1"

screen "Root screen" 800x480, template "Template_1"
   on GenerateScreen: SetTag("Tag_ScreenNumber", 1)
   TextField "HmiScreenItemData" at 1,2 size 799x54; Text 'SIEMENS NX BOTTLING ASSEMBLY LINE - HMI HOME SCREEN'
   Button "Button_1" at 113,118 size 135x57; TextOff 'START'
      on Press: SetBit("START")
      on Release: ResetBit("START")
   Button "Button_2" at 112,194 size 135x57; TextOff 'STOP'
      on Press: SetBit("STOP")
      on Release: ResetBit("STOP")
   Circle "Circle_1" at 220,123 size 23x23
      Appearance <- "CONTROL_ENABLE"
   Circle "Circle_2" at 219,198 size 22x22
      Appearance <- "CONTROL_ENABLE"
   Button "Button_3" at 300,112 size 108x40; TextOff 'Send Tall'
      on Press: SetBit("send_tall")
      on Release: ResetBit("send_tall")
   Button "Button_4" at 300,166 size 108x40; TextOff 'Send Small'
      on Press: SetBit("send_small")
      on Release: ResetBit("send_small")
   Button "Button_5" at 113,268 size 135x58; TextOff 'RESET'
      on Press: SetBit("RESET")
      on Release: ResetBit("RESET")
   Circle "Circle_3" at 220,272 size 23x23
      Appearance <- "RESTARTING"
   Circle "Circle_4" at 463,135 size 36x36
      Appearance <- "belt1"
   Circle "Circle_5" at 503,135 size 36x36
      Appearance <- "belt2_1"
   Circle "Circle_6" at 584,136 size 36x36
      Appearance <- "belt_F"
   Circle "Circle_7" at 543,135 size 36x36
      Appearance <- "belt3"
   Circle "Circle_8" at 623,136 size 36x36
      Appearance <- "belt_L"
   Circle "Circle_9" at 663,136 size 36x36
      Appearance <- "belt_R"
   TextField "Text field_1" at 472,141 size 15x23; Text '1'
   TextField "Text field_2" at 513,141 size 15x23; Text '2'
   TextField "Text field_3" at 553,141 size 15x23; Text '3'
   TextField "Text field_4" at 594,142 size 14x23; Text 'F'
   TextField "Text field_5" at 634,142 size 14x23; Text 'L'
   TextField "Text field_6" at 672,142 size 17x23; Text 'R'
   TextField "Text field_7" at 537,96 size 95x23; Text 'Belts State'
   TextField "Text field_8" at 508,203 size 158x23; Text 'ABB Robots States'
   TextField "Text field_9" at 459,249 size 81x23; Text 'ABB1 -->'
   Rectangle "Rectangle_7" at 549,248 size 74x28
      Appearance <- "ABB1_IDLE"
   Rectangle "Rectangle_8" at 632,248 size 74x28
      Appearance <- "ABB1_IDLE"
   TextField "Text field_10" at 459,296 size 81x23; Text 'ABB2 -->'
   Rectangle "Rectangle_9" at 548,295 size 74x28
      Appearance <- "ABB2_IDLE"
   Rectangle "Rectangle_10" at 631,295 size 74x28
      Appearance <- "ABB2_IDLE"
   TextField "Text field_11" at 564,251 size 43x23; Text 'IDLE'
   TextField "Text field_12" at 655,251 size 29x23; Text 'ON'
   TextField "Text field_13" at 564,298 size 43x23; Text 'IDLE'
   TextField "Text field_14" at 654,298 size 29x23; Text 'ON'
   TextField "HmiScreenItemData_1" at 1,428 size 799x51; Text 'Text'
   Button "Button_6" at 300,220 size 107x33; TextOff 'Add Cap'
      on Release: ResetBit("new_cap")
      on Press: SetBit("new_cap")
   TextField "Text field_15" at 459,343 size 78x23; Text 'Filler -->'
   Rectangle "Rectangle_14" at 548,340 size 74x30
      Appearance <- "F_FILL"
   Rectangle "Rectangle_15" at 631,339 size 73x31
      Appearance <- "F_FILL"
   TextField "Text field_16" at 562,344 size 43x23; Text 'IDLE'
   TextField "Text field_17" at 653,343 size 29x23; Text 'ON'
*)